
REGION Network 168
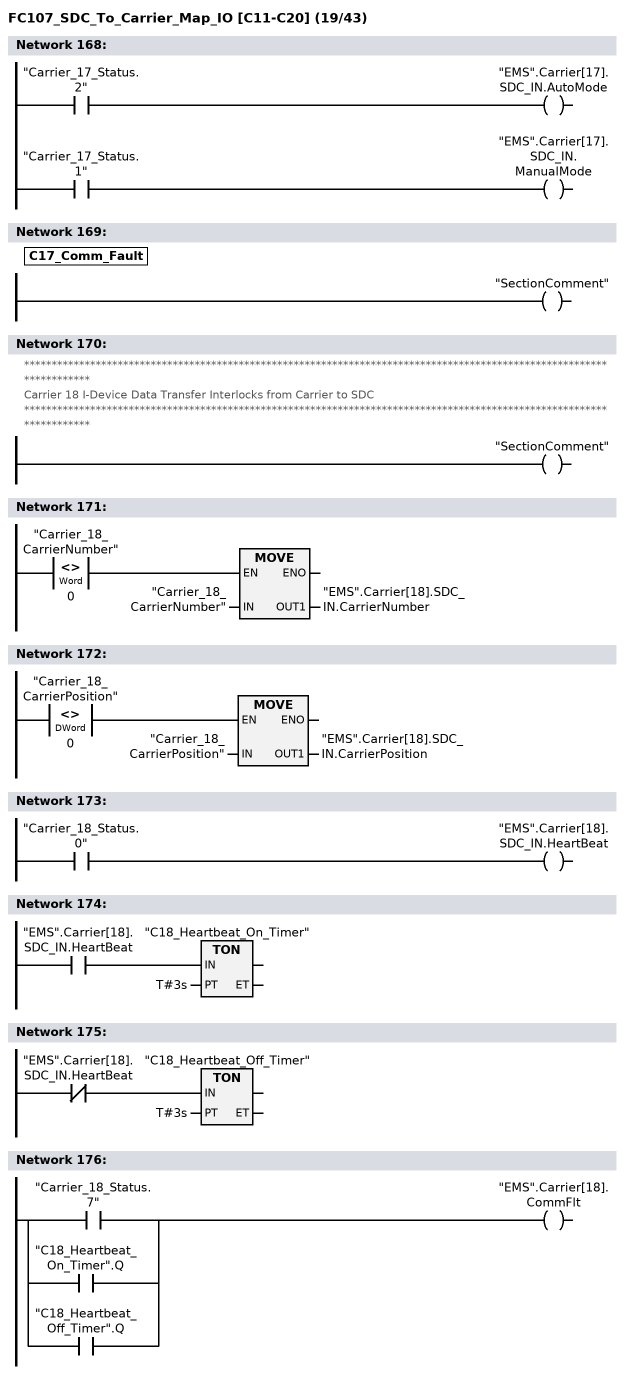
   RUNG wire#powerrail
      Contact( "Carrier_17_Status.2" )
      Coil( "EMS".Carrier[17].SDC_IN.AutoMode )
   END_RUNG
   RUNG wire#powerrail
      Contact( "Carrier_17_Status.1" )
      Coil( "EMS".Carrier[17].SDC_IN.ManualMode )
   END_RUNG
   // the same network as SCL:
   "EMS".Carrier[17].SDC_IN.AutoMode := "Carrier_17_Status.2";
   "EMS".Carrier[17].SDC_IN.ManualMode := "Carrier_17_Status.1";
END_REGION

REGION Network 169
   Label( C17_Comm_Fault )
   RUNG wire#powerrail
      Coil( "SectionComment" )
   END_RUNG
   // the same network as SCL:
   C17_Comm_Fault:
   "SectionComment" := TRUE;
END_REGION

REGION Network 170
   // **********************************************************************************************************************
   // 
   // Carrier 18 I-Device Data Transfer Interlocks from Carrier to SDC
   // 
   // **********************************************************************************************************************
   RUNG wire#powerrail
      Coil( "SectionComment" )
   END_RUNG
   // the same network as SCL:
   "SectionComment" := TRUE;
END_REGION

REGION Network 171
   RUNG wire#powerrail
      { S7_Templates := "SrcType := Word" } NE_Contact(in1 := "Carrier_18_CarrierNumber", in2 := 0)
      Move(in := "Carrier_18_CarrierNumber", out1 => "EMS".Carrier[18].SDC_IN.CarrierNumber)
   END_RUNG
   // the same network as SCL:
   IF "Carrier_18_CarrierNumber" <> 0 THEN
       "EMS".Carrier[18].SDC_IN.CarrierNumber := "Carrier_18_CarrierNumber";
   END_IF;
END_REGION

REGION Network 172
   RUNG wire#powerrail
      { S7_Templates := "SrcType := DWord" } NE_Contact(in1 := "Carrier_18_CarrierPosition", in2 := 0)
      Move(in := "Carrier_18_CarrierPosition", out1 => "EMS".Carrier[18].SDC_IN.CarrierPosition)
   END_RUNG
   // the same network as SCL:
   IF "Carrier_18_CarrierPosition" <> 0 THEN
       "EMS".Carrier[18].SDC_IN.CarrierPosition := "Carrier_18_CarrierPosition";
   END_IF;
END_REGION

REGION Network 173
   RUNG wire#powerrail
      Contact( "Carrier_18_Status.0" )
      Coil( "EMS".Carrier[18].SDC_IN.HeartBeat )
   END_RUNG
   // the same network as SCL:
   "EMS".Carrier[18].SDC_IN.HeartBeat := "Carrier_18_Status.0";
END_REGION

REGION Network 174
   "C18_Heartbeat_On_Timer".TON(IN := "EMS".Carrier[18].SDC_IN.HeartBeat, PT := T#3s);
END_REGION

REGION Network 175
   "C18_Heartbeat_Off_Timer".TON(IN := NOT "EMS".Carrier[18].SDC_IN.HeartBeat, PT := T#3s);
END_REGION

REGION Network 176
   RUNG wire#powerrail
      Contact( "Carrier_18_Status.7" )
      wire#w1
      Coil( "EMS".Carrier[18].CommFlt )
   END_RUNG
   RUNG wire#powerrail
      Contact( "C18_Heartbeat_On_Timer".Q )
   END_RUNG wire#w1
   RUNG wire#powerrail
      Contact( "C18_Heartbeat_Off_Timer".Q )
   END_RUNG wire#w1
   // the same network as SCL:
   "EMS".Carrier[18].CommFlt := "Carrier_18_Status.7" OR "C18_Heartbeat_On_Timer".Q OR "C18_Heartbeat_Off_Timer".Q;
END_REGION

REGION Network 177
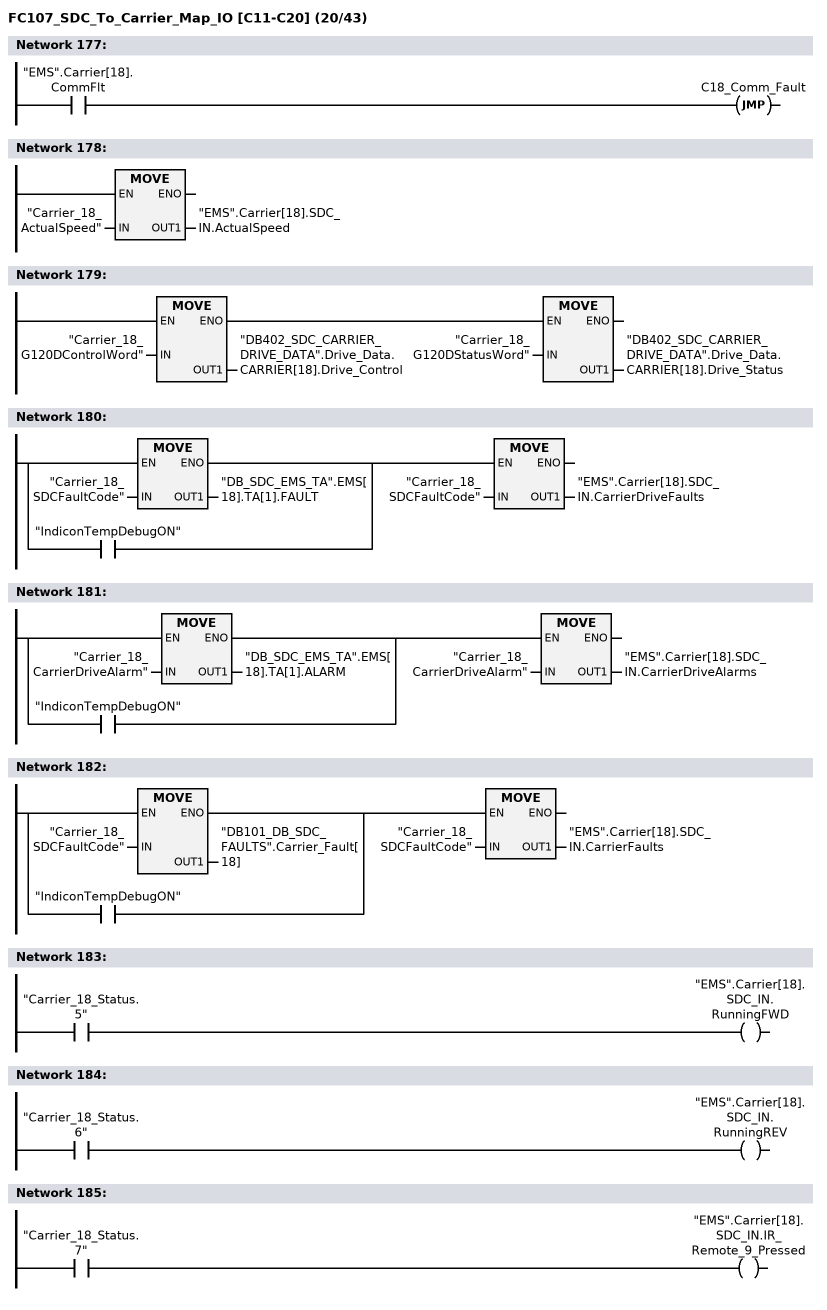
   RUNG wire#powerrail
      Contact( "EMS".Carrier[18].CommFlt )
      JumpCoil( C18_Comm_Fault )
   END_RUNG
   // the same network as SCL:
   IF "EMS".Carrier[18].CommFlt THEN GOTO C18_Comm_Fault; END_IF;
END_REGION

REGION Network 178
   RUNG wire#powerrail
      Move(in := "Carrier_18_ActualSpeed", out1 => "EMS".Carrier[18].SDC_IN.ActualSpeed)
   END_RUNG
   // the same network as SCL:
   "EMS".Carrier[18].SDC_IN.ActualSpeed := "Carrier_18_ActualSpeed";
END_REGION

REGION Network 179
   RUNG wire#powerrail
      Move(in := "Carrier_18_G120DControlWord", out1 => "DB402_SDC_CARRIER_DRIVE_DATA".Drive_Data.CARRIER[18].Drive_Control)
      Move(in := "Carrier_18_G120DStatusWord", out1 => "DB402_SDC_CARRIER_DRIVE_DATA".Drive_Data.CARRIER[18].Drive_Status)
   END_RUNG
   // the same network as SCL:
   "DB402_SDC_CARRIER_DRIVE_DATA".Drive_Data.CARRIER[18].Drive_Control := "Carrier_18_G120DControlWord";
   "DB402_SDC_CARRIER_DRIVE_DATA".Drive_Data.CARRIER[18].Drive_Status := "Carrier_18_G120DStatusWord";
END_REGION

REGION Network 180
   RUNG wire#powerrail
      Move(in := "Carrier_18_SDCFaultCode", out1 => "DB_SDC_EMS_TA".EMS[18].TA[1].FAULT)
      wire#w1
      Move(in := "Carrier_18_SDCFaultCode", out1 => "EMS".Carrier[18].SDC_IN.CarrierDriveFaults)
   END_RUNG
   RUNG wire#powerrail
      Contact( "IndiconTempDebugON" )
   END_RUNG wire#w1
   // the same network as SCL:
   "DB_SDC_EMS_TA".EMS[18].TA[1].FAULT := "Carrier_18_SDCFaultCode";
   IF TRUE OR "IndiconTempDebugON" THEN
       "EMS".Carrier[18].SDC_IN.CarrierDriveFaults := "Carrier_18_SDCFaultCode";
   END_IF;
END_REGION

REGION Network 181
   RUNG wire#powerrail
      Move(in := "Carrier_18_CarrierDriveAlarm", out1 => "DB_SDC_EMS_TA".EMS[18].TA[1].ALARM)
      wire#w1
      Move(in := "Carrier_18_CarrierDriveAlarm", out1 => "EMS".Carrier[18].SDC_IN.CarrierDriveAlarms)
   END_RUNG
   RUNG wire#powerrail
      Contact( "IndiconTempDebugON" )
   END_RUNG wire#w1
   // the same network as SCL:
   "DB_SDC_EMS_TA".EMS[18].TA[1].ALARM := "Carrier_18_CarrierDriveAlarm";
   IF TRUE OR "IndiconTempDebugON" THEN
       "EMS".Carrier[18].SDC_IN.CarrierDriveAlarms := "Carrier_18_CarrierDriveAlarm";
   END_IF;
END_REGION

REGION Network 182
   RUNG wire#powerrail
      Move(in := "Carrier_18_SDCFaultCode", out1 => "DB101_DB_SDC_FAULTS".Carrier_Fault[18])
      wire#w1
      Move(in := "Carrier_18_SDCFaultCode", out1 => "EMS".Carrier[18].SDC_IN.CarrierFaults)
   END_RUNG
   RUNG wire#powerrail
      Contact( "IndiconTempDebugON" )
   END_RUNG wire#w1
   // the same network as SCL:
   "DB101_DB_SDC_FAULTS".Carrier_Fault[18] := "Carrier_18_SDCFaultCode";
   IF TRUE OR "IndiconTempDebugON" THEN
       "EMS".Carrier[18].SDC_IN.CarrierFaults := "Carrier_18_SDCFaultCode";
   END_IF;
END_REGION

REGION Network 183
   RUNG wire#powerrail
      Contact( "Carrier_18_Status.5" )
      Coil( "EMS".Carrier[18].SDC_IN.RunningFWD )
   END_RUNG
   // the same network as SCL:
   "EMS".Carrier[18].SDC_IN.RunningFWD := "Carrier_18_Status.5";
END_REGION

REGION Network 184
   RUNG wire#powerrail
      Contact( "Carrier_18_Status.6" )
      Coil( "EMS".Carrier[18].SDC_IN.RunningREV )
   END_RUNG
   // the same network as SCL:
   "EMS".Carrier[18].SDC_IN.RunningREV := "Carrier_18_Status.6";
END_REGION

REGION Network 185
   RUNG wire#powerrail
      Contact( "Carrier_18_Status.7" )
      Coil( "EMS".Carrier[18].SDC_IN.IR_Remote_9_Pressed )
   END_RUNG
   // the same network as SCL:
   "EMS".Carrier[18].SDC_IN.IR_Remote_9_Pressed := "Carrier_18_Status.7";
END_REGION

REGION Network 186
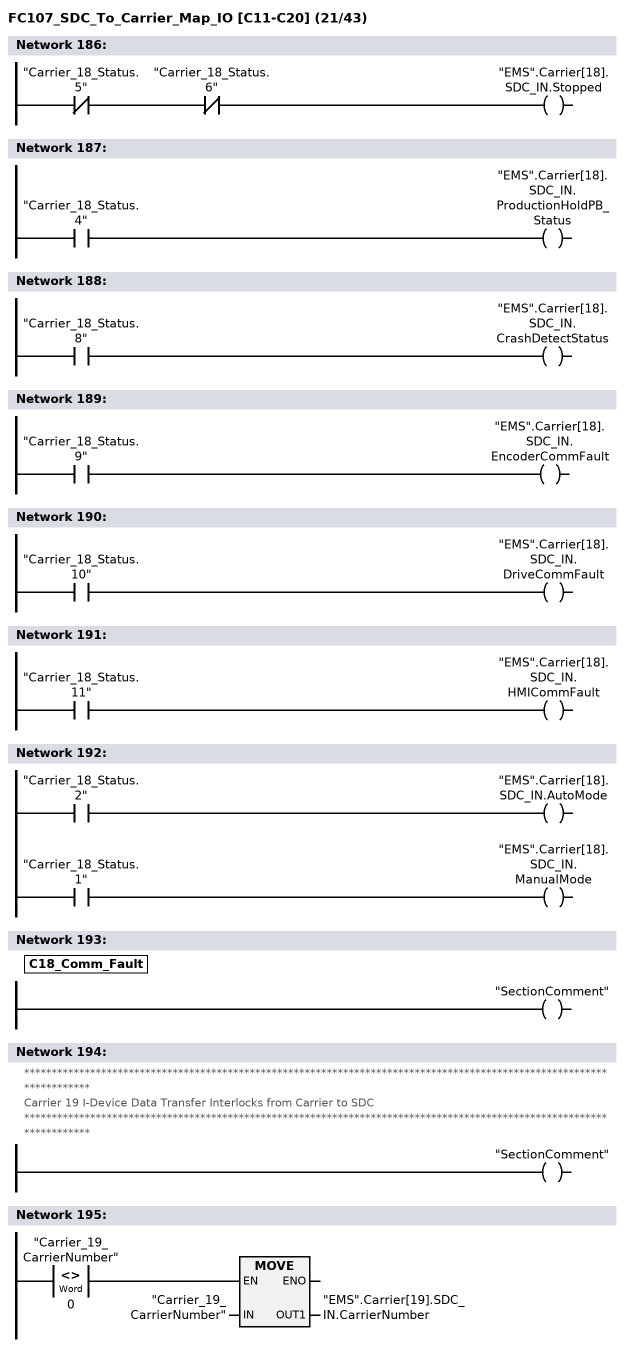
   RUNG wire#powerrail
      I_Contact( "Carrier_18_Status.5" )
      I_Contact( "Carrier_18_Status.6" )
      Coil( "EMS".Carrier[18].SDC_IN.Stopped )
   END_RUNG
   // the same network as SCL:
   "EMS".Carrier[18].SDC_IN.Stopped := NOT "Carrier_18_Status.5" AND NOT "Carrier_18_Status.6";
END_REGION

REGION Network 187
   RUNG wire#powerrail
      Contact( "Carrier_18_Status.4" )
      Coil( "EMS".Carrier[18].SDC_IN.ProductionHoldPB_Status )
   END_RUNG
   // the same network as SCL:
   "EMS".Carrier[18].SDC_IN.ProductionHoldPB_Status := "Carrier_18_Status.4";
END_REGION

REGION Network 188
   RUNG wire#powerrail
      Contact( "Carrier_18_Status.8" )
      Coil( "EMS".Carrier[18].SDC_IN.CrashDetectStatus )
   END_RUNG
   // the same network as SCL:
   "EMS".Carrier[18].SDC_IN.CrashDetectStatus := "Carrier_18_Status.8";
END_REGION

REGION Network 189
   RUNG wire#powerrail
      Contact( "Carrier_18_Status.9" )
      Coil( "EMS".Carrier[18].SDC_IN.EncoderCommFault )
   END_RUNG
   // the same network as SCL:
   "EMS".Carrier[18].SDC_IN.EncoderCommFault := "Carrier_18_Status.9";
END_REGION

REGION Network 190
   RUNG wire#powerrail
      Contact( "Carrier_18_Status.10" )
      Coil( "EMS".Carrier[18].SDC_IN.DriveCommFault )
   END_RUNG
   // the same network as SCL:
   "EMS".Carrier[18].SDC_IN.DriveCommFault := "Carrier_18_Status.10";
END_REGION

REGION Network 191
   RUNG wire#powerrail
      Contact( "Carrier_18_Status.11" )
      Coil( "EMS".Carrier[18].SDC_IN.HMICommFault )
   END_RUNG
   // the same network as SCL:
   "EMS".Carrier[18].SDC_IN.HMICommFault := "Carrier_18_Status.11";
END_REGION

REGION Network 192
   RUNG wire#powerrail
      Contact( "Carrier_18_Status.2" )
      Coil( "EMS".Carrier[18].SDC_IN.AutoMode )
   END_RUNG
   RUNG wire#powerrail
      Contact( "Carrier_18_Status.1" )
      Coil( "EMS".Carrier[18].SDC_IN.ManualMode )
   END_RUNG
   // the same network as SCL:
   "EMS".Carrier[18].SDC_IN.AutoMode := "Carrier_18_Status.2";
   "EMS".Carrier[18].SDC_IN.ManualMode := "Carrier_18_Status.1";
END_REGION

REGION Network 193
   Label( C18_Comm_Fault )
   RUNG wire#powerrail
      Coil( "SectionComment" )
   END_RUNG
   // the same network as SCL:
   C18_Comm_Fault:
   "SectionComment" := TRUE;
END_REGION

REGION Network 194
   // **********************************************************************************************************************
   // 
   // Carrier 19 I-Device Data Transfer Interlocks from Carrier to SDC
   // 
   // **********************************************************************************************************************
   RUNG wire#powerrail
      Coil( "SectionComment" )
   END_RUNG
   // the same network as SCL:
   "SectionComment" := TRUE;
END_REGION

REGION Network 195
   RUNG wire#powerrail
      { S7_Templates := "SrcType := Word" } NE_Contact(in1 := "Carrier_19_CarrierNumber", in2 := 0)
      Move(in := "Carrier_19_CarrierNumber", out1 => "EMS".Carrier[19].SDC_IN.CarrierNumber)
   END_RUNG
   // the same network as SCL:
   IF "Carrier_19_CarrierNumber" <> 0 THEN
       "EMS".Carrier[19].SDC_IN.CarrierNumber := "Carrier_19_CarrierNumber";
   END_IF;
END_REGION

REGION Network 196
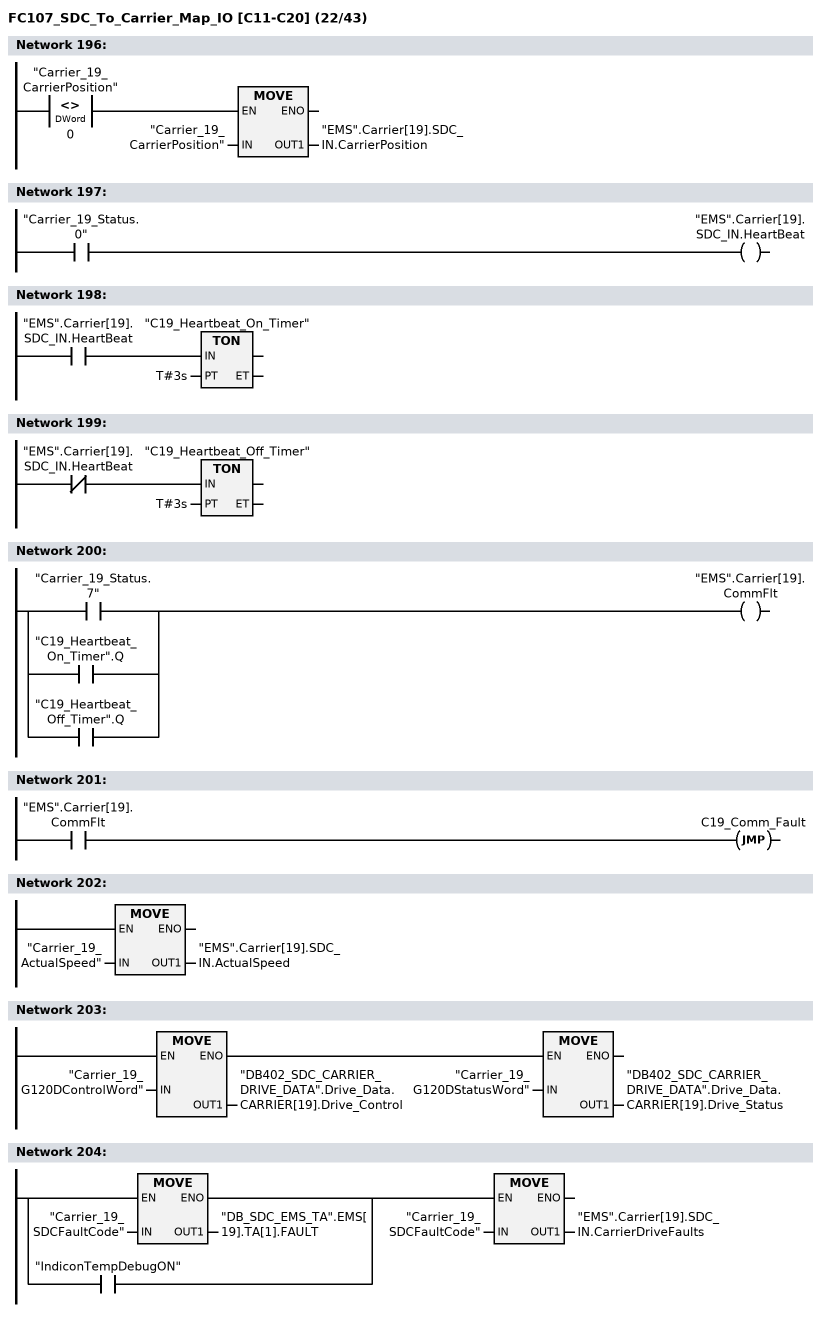
   RUNG wire#powerrail
      { S7_Templates := "SrcType := DWord" } NE_Contact(in1 := "Carrier_19_CarrierPosition", in2 := 0)
      Move(in := "Carrier_19_CarrierPosition", out1 => "EMS".Carrier[19].SDC_IN.CarrierPosition)
   END_RUNG
   // the same network as SCL:
   IF "Carrier_19_CarrierPosition" <> 0 THEN
       "EMS".Carrier[19].SDC_IN.CarrierPosition := "Carrier_19_CarrierPosition";
   END_IF;
END_REGION

REGION Network 197
   RUNG wire#powerrail
      Contact( "Carrier_19_Status.0" )
      Coil( "EMS".Carrier[19].SDC_IN.HeartBeat )
   END_RUNG
   // the same network as SCL:
   "EMS".Carrier[19].SDC_IN.HeartBeat := "Carrier_19_Status.0";
END_REGION

REGION Network 198
   "C19_Heartbeat_On_Timer".TON(IN := "EMS".Carrier[19].SDC_IN.HeartBeat, PT := T#3s);
END_REGION

REGION Network 199
   "C19_Heartbeat_Off_Timer".TON(IN := NOT "EMS".Carrier[19].SDC_IN.HeartBeat, PT := T#3s);
END_REGION

REGION Network 200
   RUNG wire#powerrail
      Contact( "Carrier_19_Status.7" )
      wire#w1
      Coil( "EMS".Carrier[19].CommFlt )
   END_RUNG
   RUNG wire#powerrail
      Contact( "C19_Heartbeat_On_Timer".Q )
   END_RUNG wire#w1
   RUNG wire#powerrail
      Contact( "C19_Heartbeat_Off_Timer".Q )
   END_RUNG wire#w1
   // the same network as SCL:
   "EMS".Carrier[19].CommFlt := "Carrier_19_Status.7" OR "C19_Heartbeat_On_Timer".Q OR "C19_Heartbeat_Off_Timer".Q;
END_REGION

REGION Network 201
   RUNG wire#powerrail
      Contact( "EMS".Carrier[19].CommFlt )
      JumpCoil( C19_Comm_Fault )
   END_RUNG
   // the same network as SCL:
   IF "EMS".Carrier[19].CommFlt THEN GOTO C19_Comm_Fault; END_IF;
END_REGION

REGION Network 202
   RUNG wire#powerrail
      Move(in := "Carrier_19_ActualSpeed", out1 => "EMS".Carrier[19].SDC_IN.ActualSpeed)
   END_RUNG
   // the same network as SCL:
   "EMS".Carrier[19].SDC_IN.ActualSpeed := "Carrier_19_ActualSpeed";
END_REGION

REGION Network 203
   RUNG wire#powerrail
      Move(in := "Carrier_19_G120DControlWord", out1 => "DB402_SDC_CARRIER_DRIVE_DATA".Drive_Data.CARRIER[19].Drive_Control)
      Move(in := "Carrier_19_G120DStatusWord", out1 => "DB402_SDC_CARRIER_DRIVE_DATA".Drive_Data.CARRIER[19].Drive_Status)
   END_RUNG
   // the same network as SCL:
   "DB402_SDC_CARRIER_DRIVE_DATA".Drive_Data.CARRIER[19].Drive_Control := "Carrier_19_G120DControlWord";
   "DB402_SDC_CARRIER_DRIVE_DATA".Drive_Data.CARRIER[19].Drive_Status := "Carrier_19_G120DStatusWord";
END_REGION

REGION Network 204
   RUNG wire#powerrail
      Move(in := "Carrier_19_SDCFaultCode", out1 => "DB_SDC_EMS_TA".EMS[19].TA[1].FAULT)
      wire#w1
      Move(in := "Carrier_19_SDCFaultCode", out1 => "EMS".Carrier[19].SDC_IN.CarrierDriveFaults)
   END_RUNG
   RUNG wire#powerrail
      Contact( "IndiconTempDebugON" )
   END_RUNG wire#w1
   // the same network as SCL:
   "DB_SDC_EMS_TA".EMS[19].TA[1].FAULT := "Carrier_19_SDCFaultCode";
   IF TRUE OR "IndiconTempDebugON" THEN
       "EMS".Carrier[19].SDC_IN.CarrierDriveFaults := "Carrier_19_SDCFaultCode";
   END_IF;
END_REGION

REGION Network 205
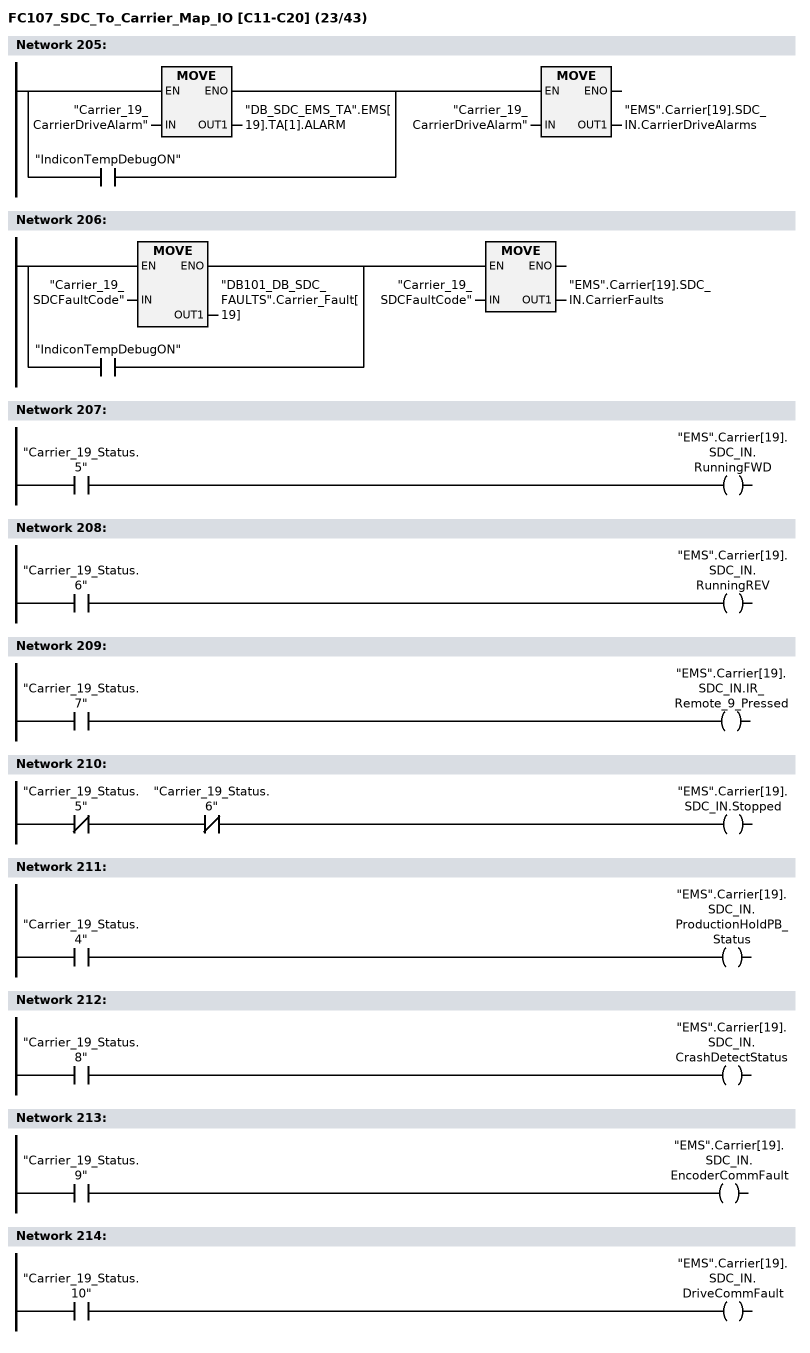
   RUNG wire#powerrail
      Move(in := "Carrier_19_CarrierDriveAlarm", out1 => "DB_SDC_EMS_TA".EMS[19].TA[1].ALARM)
      wire#w1
      Move(in := "Carrier_19_CarrierDriveAlarm", out1 => "EMS".Carrier[19].SDC_IN.CarrierDriveAlarms)
   END_RUNG
   RUNG wire#powerrail
      Contact( "IndiconTempDebugON" )
   END_RUNG wire#w1
   // the same network as SCL:
   "DB_SDC_EMS_TA".EMS[19].TA[1].ALARM := "Carrier_19_CarrierDriveAlarm";
   IF TRUE OR "IndiconTempDebugON" THEN
       "EMS".Carrier[19].SDC_IN.CarrierDriveAlarms := "Carrier_19_CarrierDriveAlarm";
   END_IF;
END_REGION

REGION Network 206
   RUNG wire#powerrail
      Move(in := "Carrier_19_SDCFaultCode", out1 => "DB101_DB_SDC_FAULTS".Carrier_Fault[19])
      wire#w1
      Move(in := "Carrier_19_SDCFaultCode", out1 => "EMS".Carrier[19].SDC_IN.CarrierFaults)
   END_RUNG
   RUNG wire#powerrail
      Contact( "IndiconTempDebugON" )
   END_RUNG wire#w1
   // the same network as SCL:
   "DB101_DB_SDC_FAULTS".Carrier_Fault[19] := "Carrier_19_SDCFaultCode";
   IF TRUE OR "IndiconTempDebugON" THEN
       "EMS".Carrier[19].SDC_IN.CarrierFaults := "Carrier_19_SDCFaultCode";
   END_IF;
END_REGION

REGION Network 207
   RUNG wire#powerrail
      Contact( "Carrier_19_Status.5" )
      Coil( "EMS".Carrier[19].SDC_IN.RunningFWD )
   END_RUNG
   // the same network as SCL:
   "EMS".Carrier[19].SDC_IN.RunningFWD := "Carrier_19_Status.5";
END_REGION

REGION Network 208
   RUNG wire#powerrail
      Contact( "Carrier_19_Status.6" )
      Coil( "EMS".Carrier[19].SDC_IN.RunningREV )
   END_RUNG
   // the same network as SCL:
   "EMS".Carrier[19].SDC_IN.RunningREV := "Carrier_19_Status.6";
END_REGION

REGION Network 209
   RUNG wire#powerrail
      Contact( "Carrier_19_Status.7" )
      Coil( "EMS".Carrier[19].SDC_IN.IR_Remote_9_Pressed )
   END_RUNG
   // the same network as SCL:
   "EMS".Carrier[19].SDC_IN.IR_Remote_9_Pressed := "Carrier_19_Status.7";
END_REGION

REGION Network 210
   RUNG wire#powerrail
      I_Contact( "Carrier_19_Status.5" )
      I_Contact( "Carrier_19_Status.6" )
      Coil( "EMS".Carrier[19].SDC_IN.Stopped )
   END_RUNG
   // the same network as SCL:
   "EMS".Carrier[19].SDC_IN.Stopped := NOT "Carrier_19_Status.5" AND NOT "Carrier_19_Status.6";
END_REGION

REGION Network 211
   RUNG wire#powerrail
      Contact( "Carrier_19_Status.4" )
      Coil( "EMS".Carrier[19].SDC_IN.ProductionHoldPB_Status )
   END_RUNG
   // the same network as SCL:
   "EMS".Carrier[19].SDC_IN.ProductionHoldPB_Status := "Carrier_19_Status.4";
END_REGION

REGION Network 212
   RUNG wire#powerrail
      Contact( "Carrier_19_Status.8" )
      Coil( "EMS".Carrier[19].SDC_IN.CrashDetectStatus )
   END_RUNG
   // the same network as SCL:
   "EMS".Carrier[19].SDC_IN.CrashDetectStatus := "Carrier_19_Status.8";
END_REGION

REGION Network 213
   RUNG wire#powerrail
      Contact( "Carrier_19_Status.9" )
      Coil( "EMS".Carrier[19].SDC_IN.EncoderCommFault )
   END_RUNG
   // the same network as SCL:
   "EMS".Carrier[19].SDC_IN.EncoderCommFault := "Carrier_19_Status.9";
END_REGION

REGION Network 214
   RUNG wire#powerrail
      Contact( "Carrier_19_Status.10" )
      Coil( "EMS".Carrier[19].SDC_IN.DriveCommFault )
   END_RUNG
   // the same network as SCL:
   "EMS".Carrier[19].SDC_IN.DriveCommFault := "Carrier_19_Status.10";
END_REGION

REGION Network 215
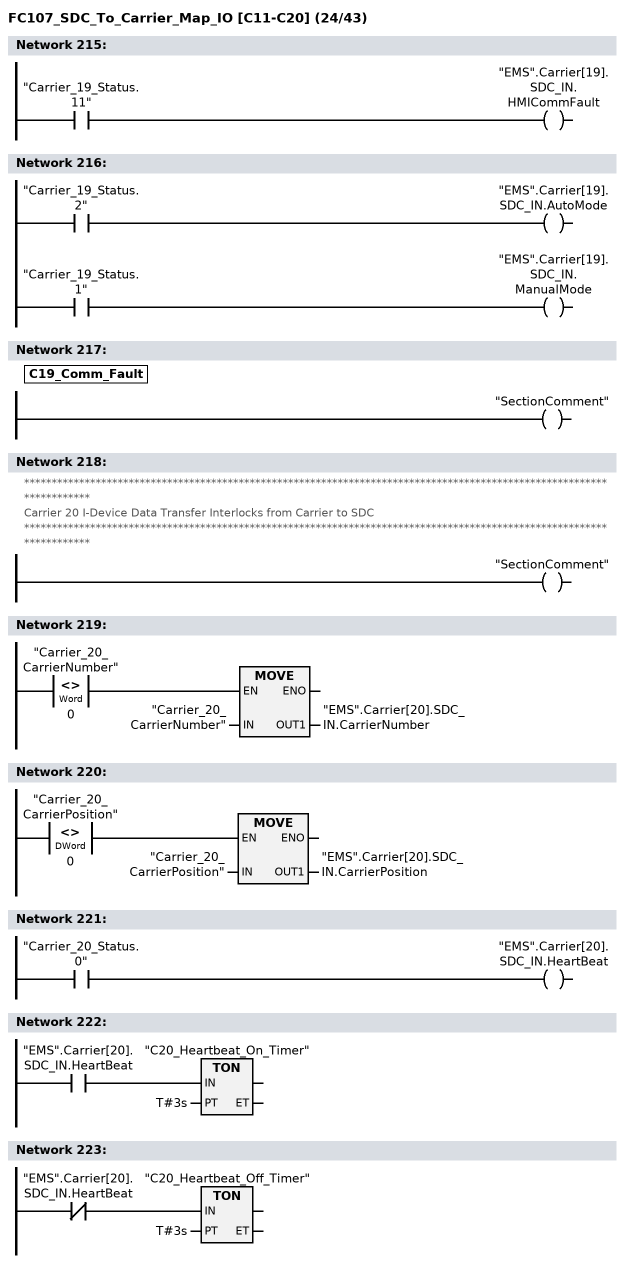
   RUNG wire#powerrail
      Contact( "Carrier_19_Status.11" )
      Coil( "EMS".Carrier[19].SDC_IN.HMICommFault )
   END_RUNG
   // the same network as SCL:
   "EMS".Carrier[19].SDC_IN.HMICommFault := "Carrier_19_Status.11";
END_REGION

REGION Network 216
   RUNG wire#powerrail
      Contact( "Carrier_19_Status.2" )
      Coil( "EMS".Carrier[19].SDC_IN.AutoMode )
   END_RUNG
   RUNG wire#powerrail
      Contact( "Carrier_19_Status.1" )
      Coil( "EMS".Carrier[19].SDC_IN.ManualMode )
   END_RUNG
   // the same network as SCL:
   "EMS".Carrier[19].SDC_IN.AutoMode := "Carrier_19_Status.2";
   "EMS".Carrier[19].SDC_IN.ManualMode := "Carrier_19_Status.1";
END_REGION

REGION Network 217
   Label( C19_Comm_Fault )
   RUNG wire#powerrail
      Coil( "SectionComment" )
   END_RUNG
   // the same network as SCL:
   C19_Comm_Fault:
   "SectionComment" := TRUE;
END_REGION

REGION Network 218
   // **********************************************************************************************************************
   // 
   // Carrier 20 I-Device Data Transfer Interlocks from Carrier to SDC
   // 
   // **********************************************************************************************************************
   RUNG wire#powerrail
      Coil( "SectionComment" )
   END_RUNG
   // the same network as SCL:
   "SectionComment" := TRUE;
END_REGION

REGION Network 219
   RUNG wire#powerrail
      { S7_Templates := "SrcType := Word" } NE_Contact(in1 := "Carrier_20_CarrierNumber", in2 := 0)
      Move(in := "Carrier_20_CarrierNumber", out1 => "EMS".Carrier[20].SDC_IN.CarrierNumber)
   END_RUNG
   // the same network as SCL:
   IF "Carrier_20_CarrierNumber" <> 0 THEN
       "EMS".Carrier[20].SDC_IN.CarrierNumber := "Carrier_20_CarrierNumber";
   END_IF;
END_REGION

REGION Network 220
   RUNG wire#powerrail
      { S7_Templates := "SrcType := DWord" } NE_Contact(in1 := "Carrier_20_CarrierPosition", in2 := 0)
      Move(in := "Carrier_20_CarrierPosition", out1 => "EMS".Carrier[20].SDC_IN.CarrierPosition)
   END_RUNG
   // the same network as SCL:
   IF "Carrier_20_CarrierPosition" <> 0 THEN
       "EMS".Carrier[20].SDC_IN.CarrierPosition := "Carrier_20_CarrierPosition";
   END_IF;
END_REGION

REGION Network 221
   RUNG wire#powerrail
      Contact( "Carrier_20_Status.0" )
      Coil( "EMS".Carrier[20].SDC_IN.HeartBeat )
   END_RUNG
   // the same network as SCL:
   "EMS".Carrier[20].SDC_IN.HeartBeat := "Carrier_20_Status.0";
END_REGION

REGION Network 222
   "C20_Heartbeat_On_Timer".TON(IN := "EMS".Carrier[20].SDC_IN.HeartBeat, PT := T#3s);
END_REGION

REGION Network 223
   "C20_Heartbeat_Off_Timer".TON(IN := NOT "EMS".Carrier[20].SDC_IN.HeartBeat, PT := T#3s);
END_REGION

REGION Network 224
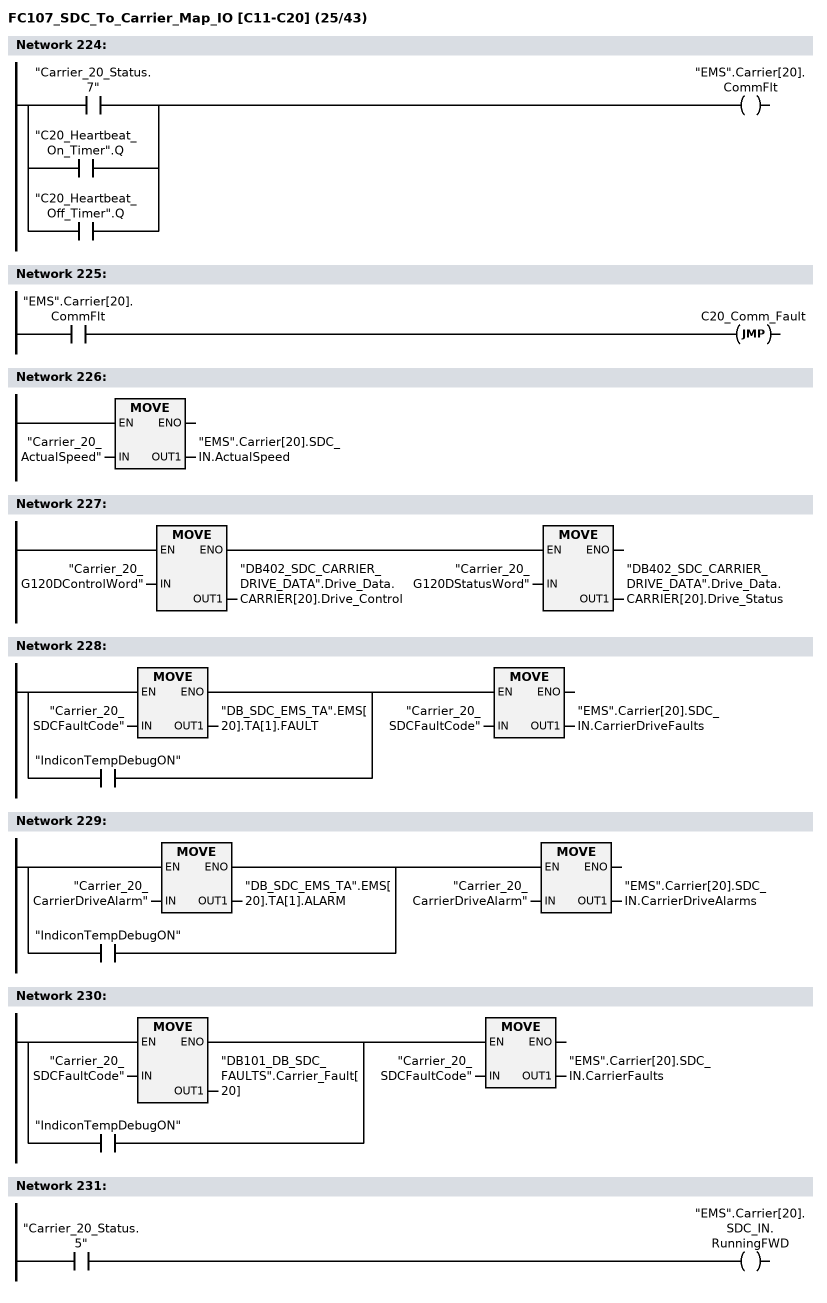
   RUNG wire#powerrail
      Contact( "Carrier_20_Status.7" )
      wire#w1
      Coil( "EMS".Carrier[20].CommFlt )
   END_RUNG
   RUNG wire#powerrail
      Contact( "C20_Heartbeat_On_Timer".Q )
   END_RUNG wire#w1
   RUNG wire#powerrail
      Contact( "C20_Heartbeat_Off_Timer".Q )
   END_RUNG wire#w1
   // the same network as SCL:
   "EMS".Carrier[20].CommFlt := "Carrier_20_Status.7" OR "C20_Heartbeat_On_Timer".Q OR "C20_Heartbeat_Off_Timer".Q;
END_REGION

REGION Network 225
   RUNG wire#powerrail
      Contact( "EMS".Carrier[20].CommFlt )
      JumpCoil( C20_Comm_Fault )
   END_RUNG
   // the same network as SCL:
   IF "EMS".Carrier[20].CommFlt THEN GOTO C20_Comm_Fault; END_IF;
END_REGION

REGION Network 226
   RUNG wire#powerrail
      Move(in := "Carrier_20_ActualSpeed", out1 => "EMS".Carrier[20].SDC_IN.ActualSpeed)
   END_RUNG
   // the same network as SCL:
   "EMS".Carrier[20].SDC_IN.ActualSpeed := "Carrier_20_ActualSpeed";
END_REGION

REGION Network 227
   RUNG wire#powerrail
      Move(in := "Carrier_20_G120DControlWord", out1 => "DB402_SDC_CARRIER_DRIVE_DATA".Drive_Data.CARRIER[20].Drive_Control)
      Move(in := "Carrier_20_G120DStatusWord", out1 => "DB402_SDC_CARRIER_DRIVE_DATA".Drive_Data.CARRIER[20].Drive_Status)
   END_RUNG
   // the same network as SCL:
   "DB402_SDC_CARRIER_DRIVE_DATA".Drive_Data.CARRIER[20].Drive_Control := "Carrier_20_G120DControlWord";
   "DB402_SDC_CARRIER_DRIVE_DATA".Drive_Data.CARRIER[20].Drive_Status := "Carrier_20_G120DStatusWord";
END_REGION

REGION Network 228
   RUNG wire#powerrail
      Move(in := "Carrier_20_SDCFaultCode", out1 => "DB_SDC_EMS_TA".EMS[20].TA[1].FAULT)
      wire#w1
      Move(in := "Carrier_20_SDCFaultCode", out1 => "EMS".Carrier[20].SDC_IN.CarrierDriveFaults)
   END_RUNG
   RUNG wire#powerrail
      Contact( "IndiconTempDebugON" )
   END_RUNG wire#w1
   // the same network as SCL:
   "DB_SDC_EMS_TA".EMS[20].TA[1].FAULT := "Carrier_20_SDCFaultCode";
   IF TRUE OR "IndiconTempDebugON" THEN
       "EMS".Carrier[20].SDC_IN.CarrierDriveFaults := "Carrier_20_SDCFaultCode";
   END_IF;
END_REGION

REGION Network 229
   RUNG wire#powerrail
      Move(in := "Carrier_20_CarrierDriveAlarm", out1 => "DB_SDC_EMS_TA".EMS[20].TA[1].ALARM)
      wire#w1
      Move(in := "Carrier_20_CarrierDriveAlarm", out1 => "EMS".Carrier[20].SDC_IN.CarrierDriveAlarms)
   END_RUNG
   RUNG wire#powerrail
      Contact( "IndiconTempDebugON" )
   END_RUNG wire#w1
   // the same network as SCL:
   "DB_SDC_EMS_TA".EMS[20].TA[1].ALARM := "Carrier_20_CarrierDriveAlarm";
   IF TRUE OR "IndiconTempDebugON" THEN
       "EMS".Carrier[20].SDC_IN.CarrierDriveAlarms := "Carrier_20_CarrierDriveAlarm";
   END_IF;
END_REGION

REGION Network 230
   RUNG wire#powerrail
      Move(in := "Carrier_20_SDCFaultCode", out1 => "DB101_DB_SDC_FAULTS".Carrier_Fault[20])
      wire#w1
      Move(in := "Carrier_20_SDCFaultCode", out1 => "EMS".Carrier[20].SDC_IN.CarrierFaults)
   END_RUNG
   RUNG wire#powerrail
      Contact( "IndiconTempDebugON" )
   END_RUNG wire#w1
   // the same network as SCL:
   "DB101_DB_SDC_FAULTS".Carrier_Fault[20] := "Carrier_20_SDCFaultCode";
   IF TRUE OR "IndiconTempDebugON" THEN
       "EMS".Carrier[20].SDC_IN.CarrierFaults := "Carrier_20_SDCFaultCode";
   END_IF;
END_REGION

REGION Network 231
   RUNG wire#powerrail
      Contact( "Carrier_20_Status.5" )
      Coil( "EMS".Carrier[20].SDC_IN.RunningFWD )
   END_RUNG
   // the same network as SCL:
   "EMS".Carrier[20].SDC_IN.RunningFWD := "Carrier_20_Status.5";
END_REGION

REGION Network 232
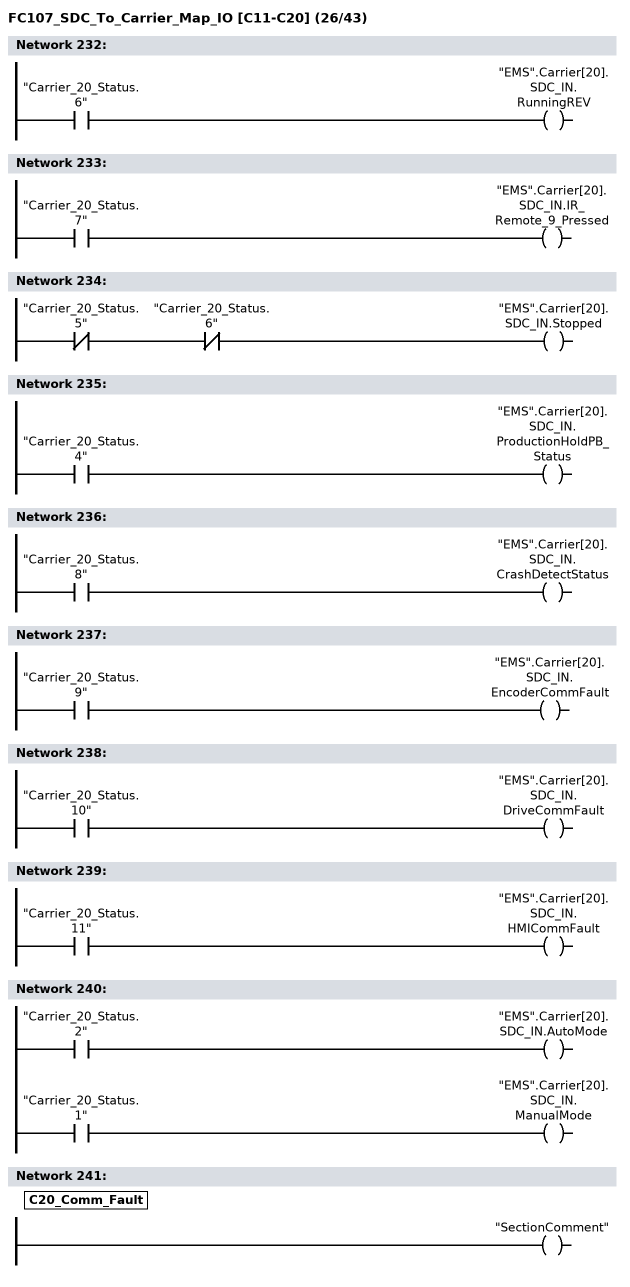
   RUNG wire#powerrail
      Contact( "Carrier_20_Status.6" )
      Coil( "EMS".Carrier[20].SDC_IN.RunningREV )
   END_RUNG
   // the same network as SCL:
   "EMS".Carrier[20].SDC_IN.RunningREV := "Carrier_20_Status.6";
END_REGION

REGION Network 233
   RUNG wire#powerrail
      Contact( "Carrier_20_Status.7" )
      Coil( "EMS".Carrier[20].SDC_IN.IR_Remote_9_Pressed )
   END_RUNG
   // the same network as SCL:
   "EMS".Carrier[20].SDC_IN.IR_Remote_9_Pressed := "Carrier_20_Status.7";
END_REGION

REGION Network 234
   RUNG wire#powerrail
      I_Contact( "Carrier_20_Status.5" )
      I_Contact( "Carrier_20_Status.6" )
      Coil( "EMS".Carrier[20].SDC_IN.Stopped )
   END_RUNG
   // the same network as SCL:
   "EMS".Carrier[20].SDC_IN.Stopped := NOT "Carrier_20_Status.5" AND NOT "Carrier_20_Status.6";
END_REGION

REGION Network 235
   RUNG wire#powerrail
      Contact( "Carrier_20_Status.4" )
      Coil( "EMS".Carrier[20].SDC_IN.ProductionHoldPB_Status )
   END_RUNG
   // the same network as SCL:
   "EMS".Carrier[20].SDC_IN.ProductionHoldPB_Status := "Carrier_20_Status.4";
END_REGION

REGION Network 236
   RUNG wire#powerrail
      Contact( "Carrier_20_Status.8" )
      Coil( "EMS".Carrier[20].SDC_IN.CrashDetectStatus )
   END_RUNG
   // the same network as SCL:
   "EMS".Carrier[20].SDC_IN.CrashDetectStatus := "Carrier_20_Status.8";
END_REGION

REGION Network 237
   RUNG wire#powerrail
      Contact( "Carrier_20_Status.9" )
      Coil( "EMS".Carrier[20].SDC_IN.EncoderCommFault )
   END_RUNG
   // the same network as SCL:
   "EMS".Carrier[20].SDC_IN.EncoderCommFault := "Carrier_20_Status.9";
END_REGION

REGION Network 238
   RUNG wire#powerrail
      Contact( "Carrier_20_Status.10" )
      Coil( "EMS".Carrier[20].SDC_IN.DriveCommFault )
   END_RUNG
   // the same network as SCL:
   "EMS".Carrier[20].SDC_IN.DriveCommFault := "Carrier_20_Status.10";
END_REGION

REGION Network 239
   RUNG wire#powerrail
      Contact( "Carrier_20_Status.11" )
      Coil( "EMS".Carrier[20].SDC_IN.HMICommFault )
   END_RUNG
   // the same network as SCL:
   "EMS".Carrier[20].SDC_IN.HMICommFault := "Carrier_20_Status.11";
END_REGION

REGION Network 240
   RUNG wire#powerrail
      Contact( "Carrier_20_Status.2" )
      Coil( "EMS".Carrier[20].SDC_IN.AutoMode )
   END_RUNG
   RUNG wire#powerrail
      Contact( "Carrier_20_Status.1" )
      Coil( "EMS".Carrier[20].SDC_IN.ManualMode )
   END_RUNG
   // the same network as SCL:
   "EMS".Carrier[20].SDC_IN.AutoMode := "Carrier_20_Status.2";
   "EMS".Carrier[20].SDC_IN.ManualMode := "Carrier_20_Status.1";
END_REGION

REGION Network 241
   Label( C20_Comm_Fault )
   RUNG wire#powerrail
      Coil( "SectionComment" )
   END_RUNG
   // the same network as SCL:
   C20_Comm_Fault:
   "SectionComment" := TRUE;
END_REGION

REGION Network 242
